(* Logix 5000 project; controller PLC_MCC1201_220AP1 vendor 1 type 14 code 164 rev 35.11; software revision 35.00; part 22 of 25 *)
(* tags used below, declared in another part *)
   LEHR_dActualSpeedValue_mm_min : DINT;
   LEHR_dLehrPositionAdvancement : DINT;
   TMP_dDistanceBetweenCut : DINT;
   TMP_xSimulationMode : BOOL;
   DISTANCE : ALIAS FOR N7[1];
   M203DROP_HMR : MAC_DROPCONV_HMR;
   M225 : MAC_EMERGENCYXCUT;
   M225_ALM : MAC_EMERGENCYXCUT_ALM;
   M225_HMR : MAC_EMERGENCYXCUT_HMR;
   M225_HMW : MAC_EMERGENCYXCUT_HMW;
   M225_IN_MOTION : MAC_EMERGENCYXCUT_IN_MOTION;
   M225_M1_DR : AXIS_CIP_DRIVE;
   M225_OUT_MOTION : MAC_EMERGENCYXCUT_OUT_MOTION;
   N54 : DINT[501];
   Status : INT;   // INT tag to retrieve Status value through GSV created during conversion
   TMP_dIndex : DINT;
   Z200_UPS : ZONE_UPS;
(* MainProgram, continued *)

ROUTINE M225_EmCut_Faults   (* ladder *)
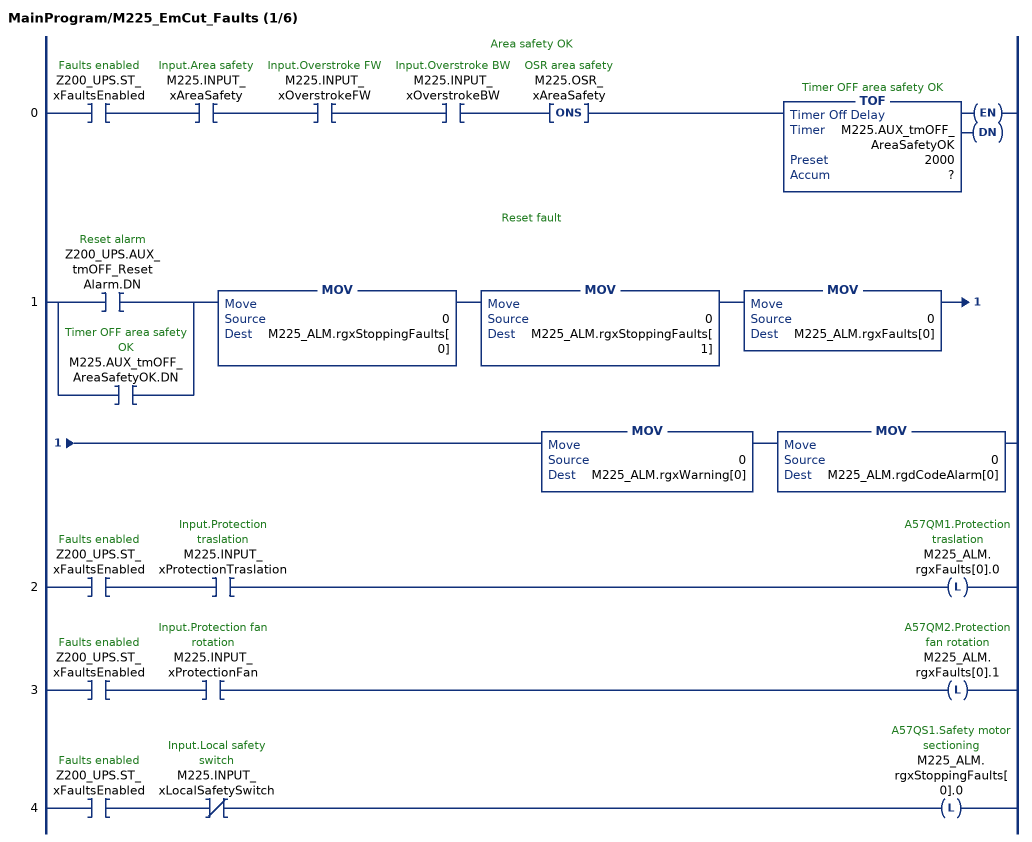
   // Area safety OK
   0: XIC(Z200_UPS.ST_xFaultsEnabled)XIC(M225.INPUT_xAreaSafety)XIC(M225.INPUT_xOverstrokeFW)XIC(M225.INPUT_xOverstrokeBW)ONS(M225.OSR_xAreaSafety)TOF(M225.AUX_tmOFF_AreaSafetyOK,?,?);
   // Reset fault
   1: [XIC(Z200_UPS.AUX_tmOFF_ResetAlarm.DN) ,XIC(M225.AUX_tmOFF_AreaSafetyOK.DN) ]MOV(0,M225_ALM.rgxStoppingFaults[0])MOV(0,M225_ALM.rgxStoppingFaults[1])MOV(0,M225_ALM.rgxFaults[0])MOV(0,M225_ALM.rgxWarning[0])MOV(0,M225_ALM.rgdCodeAlarm[0]);
   2: XIC(Z200_UPS.ST_xFaultsEnabled)XIC(M225.INPUT_xProtectionTraslation)OTL(M225_ALM.rgxFaults[0].0);
   3: XIC(Z200_UPS.ST_xFaultsEnabled)XIC(M225.INPUT_xProtectionFan)OTL(M225_ALM.rgxFaults[0].1);
   4: XIC(Z200_UPS.ST_xFaultsEnabled)XIO(M225.INPUT_xLocalSafetySwitch)OTL(M225_ALM.rgxStoppingFaults[0].0);
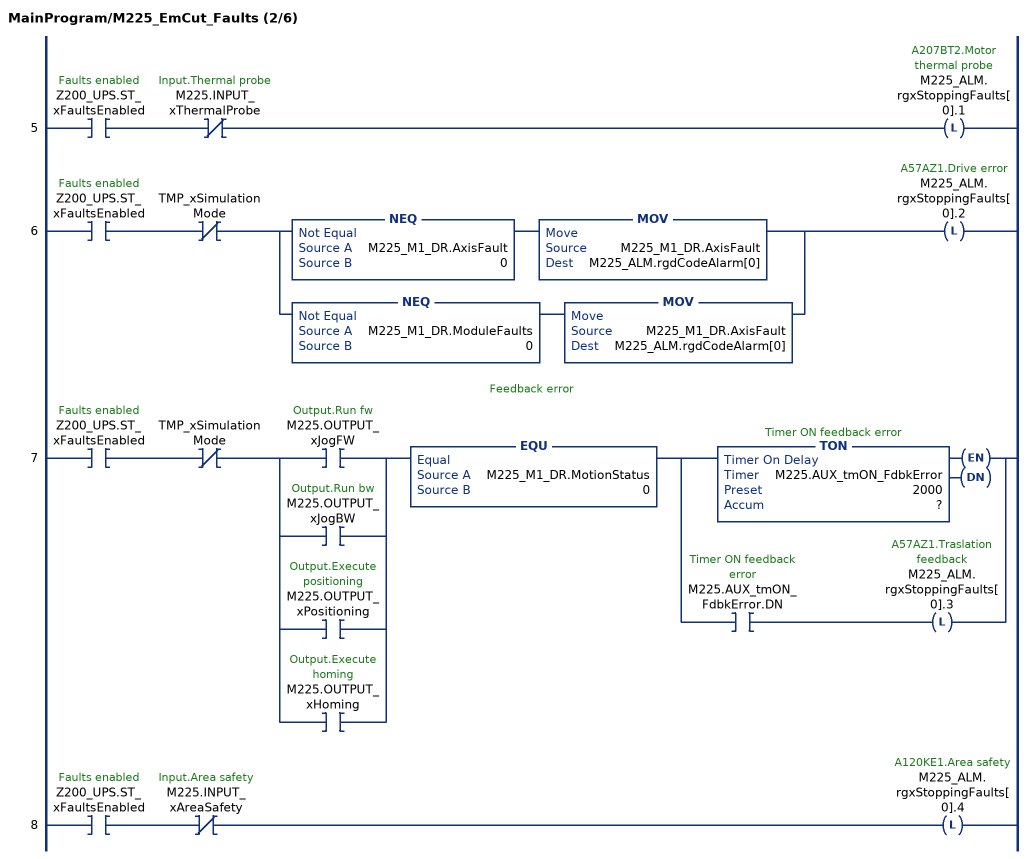
   5: XIC(Z200_UPS.ST_xFaultsEnabled)XIO(M225.INPUT_xThermalProbe)OTL(M225_ALM.rgxStoppingFaults[0].1);
   6: XIC(Z200_UPS.ST_xFaultsEnabled)XIO(TMP_xSimulationMode)[NEQ(M225_M1_DR.AxisFault,0) MOV(M225_M1_DR.AxisFault,M225_ALM.rgdCodeAlarm[0]) ,NEQ(M225_M1_DR.ModuleFaults,0) MOV(M225_M1_DR.AxisFault,M225_ALM.rgdCodeAlarm[0]) ]OTL(M225_ALM.rgxStoppingFaults[0].2);
   // Feedback error
   7: XIC(Z200_UPS.ST_xFaultsEnabled)XIO(TMP_xSimulationMode)[XIC(M225.OUTPUT_xJogFW) ,XIC(M225.OUTPUT_xJogBW) ,XIC(M225.OUTPUT_xPositioning) ,XIC(M225.OUTPUT_xHoming) ]EQU(M225_M1_DR.MotionStatus,0)[TON(M225.AUX_tmON_FdbkError,?,?) ,XIC(M225.AUX_tmON_FdbkError.DN) OTL(M225_ALM.rgxStoppingFaults[0].3) ];
   8: XIC(Z200_UPS.ST_xFaultsEnabled)XIO(M225.INPUT_xAreaSafety)OTL(M225_ALM.rgxStoppingFaults[0].4);
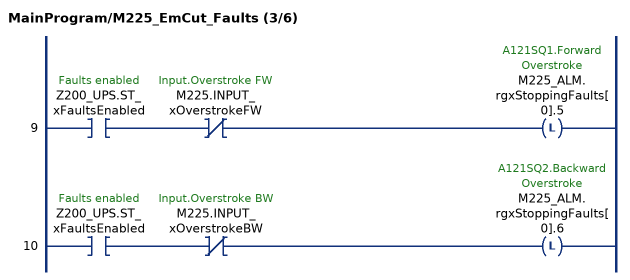
   9: XIC(Z200_UPS.ST_xFaultsEnabled)XIO(M225.INPUT_xOverstrokeFW)OTL(M225_ALM.rgxStoppingFaults[0].5);
   10: XIC(Z200_UPS.ST_xFaultsEnabled)XIO(M225.INPUT_xOverstrokeBW)OTL(M225_ALM.rgxStoppingFaults[0].6);
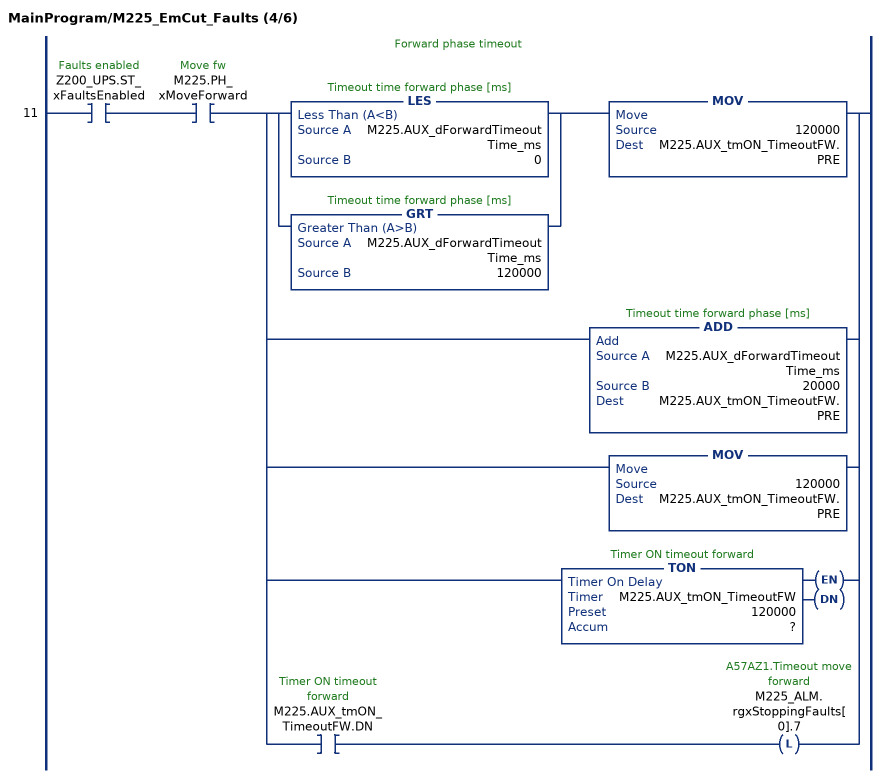
   // Forward phase timeout
   11: XIC(Z200_UPS.ST_xFaultsEnabled)XIC(M225.PH_xMoveForward)[[LES(M225.AUX_dForwardTimeoutTime_ms,0) ,GRT(M225.AUX_dForwardTimeoutTime_ms,120000) ] MOV(120000,M225.AUX_tmON_TimeoutFW.PRE) ,ADD(M225.AUX_dForwardTimeoutTime_ms,20000,M225.AUX_tmON_TimeoutFW.PRE) ,MOV(120000,M225.AUX_tmON_TimeoutFW.PRE) ,TON(M225.AUX_tmON_TimeoutFW,?,?) ,XIC(M225.AUX_tmON_TimeoutFW.DN) OTL(M225_ALM.rgxStoppingFaults[0].7) ];
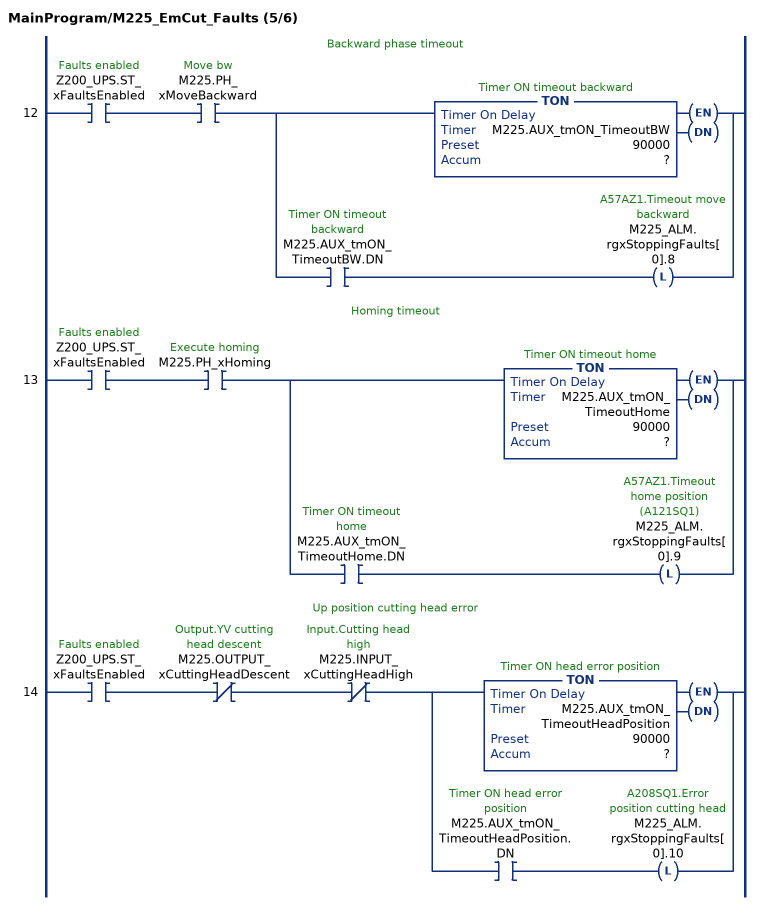
   // Backward phase timeout
   12: XIC(Z200_UPS.ST_xFaultsEnabled)XIC(M225.PH_xMoveBackward)[TON(M225.AUX_tmON_TimeoutBW,?,?) ,XIC(M225.AUX_tmON_TimeoutBW.DN) OTL(M225_ALM.rgxStoppingFaults[0].8) ];
   // Homing timeout
   13: XIC(Z200_UPS.ST_xFaultsEnabled)XIC(M225.PH_xHoming)[TON(M225.AUX_tmON_TimeoutHome,?,?) ,XIC(M225.AUX_tmON_TimeoutHome.DN) OTL(M225_ALM.rgxStoppingFaults[0].9) ];
   // Up position cutting head error
   14: XIC(Z200_UPS.ST_xFaultsEnabled)XIO(M225.OUTPUT_xCuttingHeadDescent)XIO(M225.INPUT_xCuttingHeadHigh)[TON(M225.AUX_tmON_TimeoutHeadPosition,?,?) ,XIC(M225.AUX_tmON_TimeoutHeadPosition.DN) OTL(M225_ALM.rgxStoppingFaults[0].10) ];
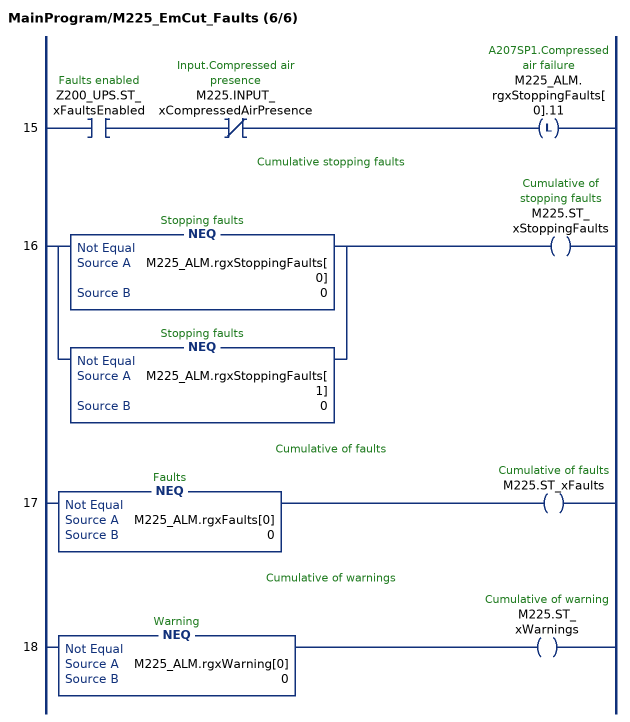
   15: XIC(Z200_UPS.ST_xFaultsEnabled)XIO(M225.INPUT_xCompressedAirPresence)OTL(M225_ALM.rgxStoppingFaults[0].11);
   // Cumulative stopping faults
   16: [NEQ(M225_ALM.rgxStoppingFaults[0],0) ,NEQ(M225_ALM.rgxStoppingFaults[1],0) ]OTE(M225.ST_xStoppingFaults);
   // Cumulative of faults
   17: NEQ(M225_ALM.rgxFaults[0],0)OTE(M225.ST_xFaults);
   // Cumulative of warnings
   18: NEQ(M225_ALM.rgxWarning[0],0)OTE(M225.ST_xWarnings);
END_ROUTINE

ROUTINE M225_EmCut_FIFOTank   (* structured text *)
   FOR TMP_dIndex:=0 TO M225.AUX_dTankElementCounter-1 DO
   	M225.AUX_rgdCutTank[TMP_dIndex]:=M225.AUX_rgdCutTank[TMP_dIndex+1];
   END_FOR;
END_ROUTINE

ROUTINE M225_EmCut_Logics   (* ladder *)
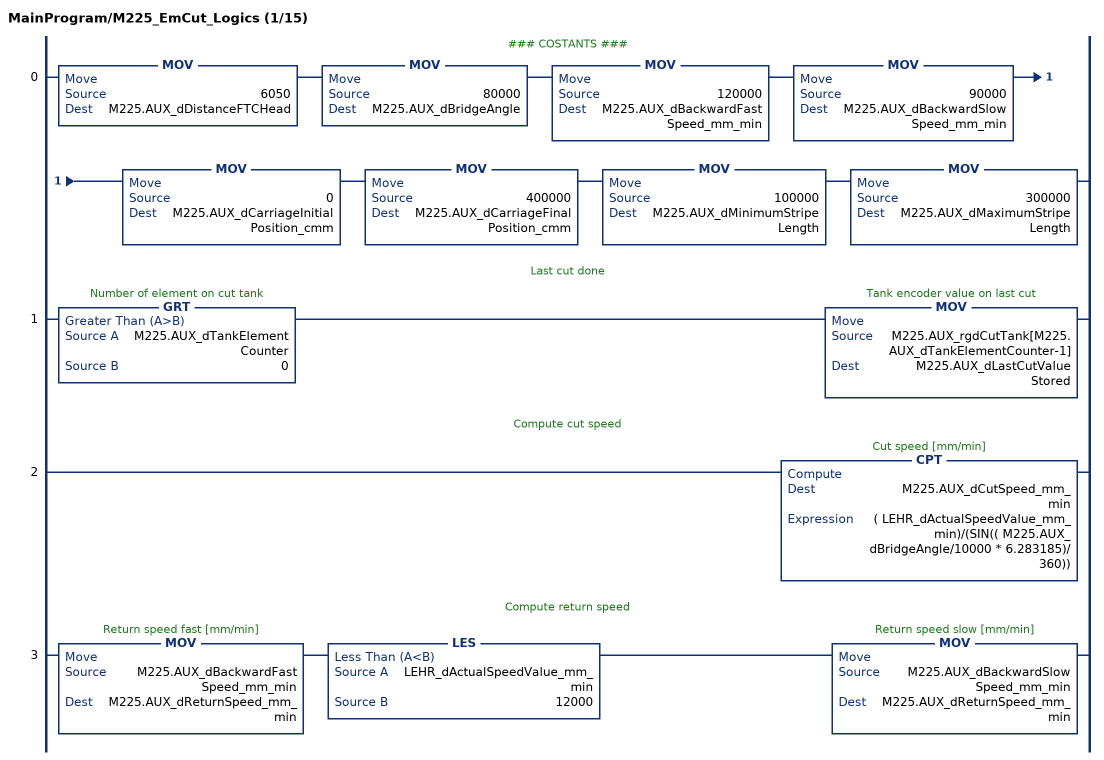
   // ### COSTANTS ###
   0: MOV(6050,M225.AUX_dDistanceFTCHead)MOV(80000,M225.AUX_dBridgeAngle)MOV(120000,M225.AUX_dBackwardFastSpeed_mm_min)MOV(90000,M225.AUX_dBackwardSlowSpeed_mm_min)MOV(0,M225.AUX_dCarriageInitialPosition_cmm)MOV(400000,M225.AUX_dCarriageFinalPosition_cmm)MOV(100000,M225.AUX_dMinimumStripeLength)MOV(300000,M225.AUX_dMaximumStripeLength);
   // Last cut done
   1: GRT(M225.AUX_dTankElementCounter,0)MOV(M225.AUX_rgdCutTank[M225.AUX_dTankElementCounter-1],M225.AUX_dLastCutValueStored);
   // Compute cut speed
   2: CPT(M225.AUX_dCutSpeed_mm_min,( LEHR_dActualSpeedValue_mm_min)/(SIN(( M225.AUX_dBridgeAngle/10000 * 6.283185)/ 360)));
   // Compute return speed
   3: MOV(M225.AUX_dBackwardFastSpeed_mm_min,M225.AUX_dReturnSpeed_mm_min)LES(LEHR_dActualSpeedValue_mm_min,12000)MOV(M225.AUX_dBackwardSlowSpeed_mm_min,M225.AUX_dReturnSpeed_mm_min);
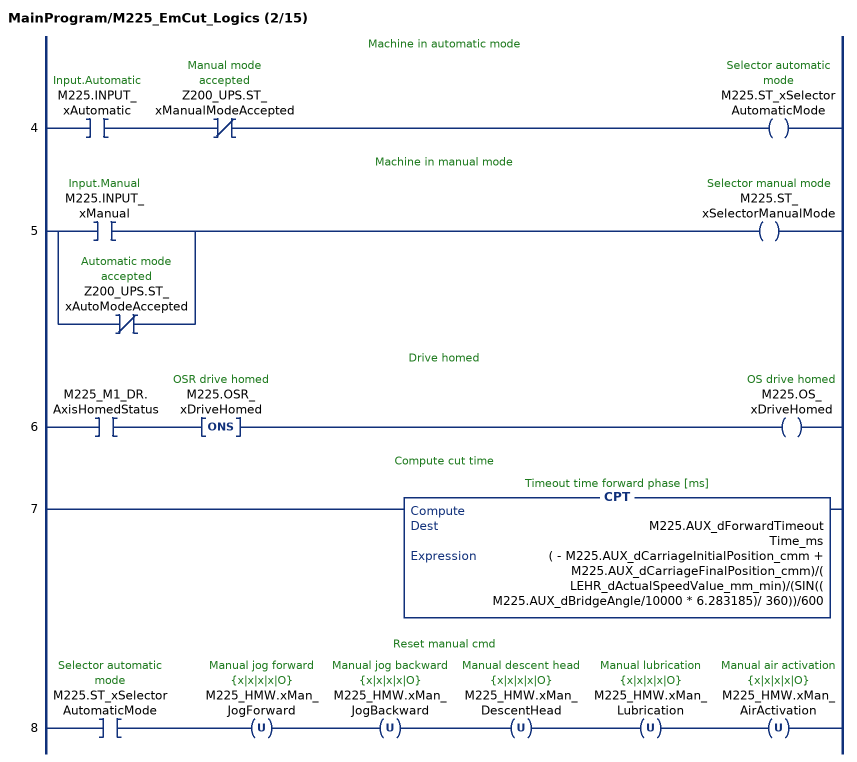
   // Machine in automatic mode
   4: XIC(M225.INPUT_xAutomatic)XIO(Z200_UPS.ST_xManualModeAccepted)OTE(M225.ST_xSelectorAutomaticMode);
   // Machine in manual mode
   5: [XIC(M225.INPUT_xManual) ,XIO(Z200_UPS.ST_xAutoModeAccepted) ]OTE(M225.ST_xSelectorManualMode);
   // Drive homed
   6: XIC(M225_M1_DR.AxisHomedStatus)ONS(M225.OSR_xDriveHomed)OTE(M225.OS_xDriveHomed);
   // Compute cut time
   7: CPT(M225.AUX_dForwardTimeoutTime_ms,( - M225.AUX_dCarriageInitialPosition_cmm + M225.AUX_dCarriageFinalPosition_cmm)/( LEHR_dActualSpeedValue_mm_min)/(SIN(( M225.AUX_dBridgeAngle/10000 * 6.283185)/ 360))/600);
   // Reset manual cmd
   8: XIC(M225.ST_xSelectorAutomaticMode)OTU(M225_HMW.xMan_JogForward)OTU(M225_HMW.xMan_JogBackward)OTU(M225_HMW.xMan_DescentHead)OTU(M225_HMW.xMan_Lubrication)OTU(M225_HMW.xMan_AirActivation);
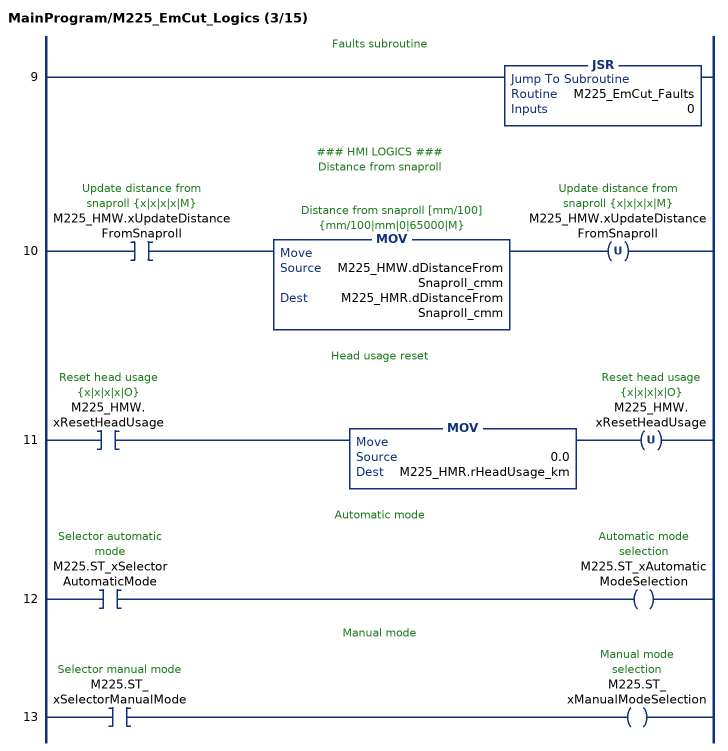
   // Faults subroutine
   9: JSR(M225_EmCut_Faults,0);
   // ### HMI LOGICS ###
   // Distance from snaproll
   10: XIC(M225_HMW.xUpdateDistanceFromSnaproll)MOV(M225_HMW.dDistanceFromSnaproll_cmm,M225_HMR.dDistanceFromSnaproll_cmm)OTU(M225_HMW.xUpdateDistanceFromSnaproll);
   // Head usage reset
   11: XIC(M225_HMW.xResetHeadUsage)MOV(0.0,M225_HMR.rHeadUsage_km)OTU(M225_HMW.xResetHeadUsage);
   // Automatic mode
   12: XIC(M225.ST_xSelectorAutomaticMode)OTE(M225.ST_xAutomaticModeSelection);
   // Manual mode
   13: XIC(M225.ST_xSelectorManualMode)OTE(M225.ST_xManualModeSelection);
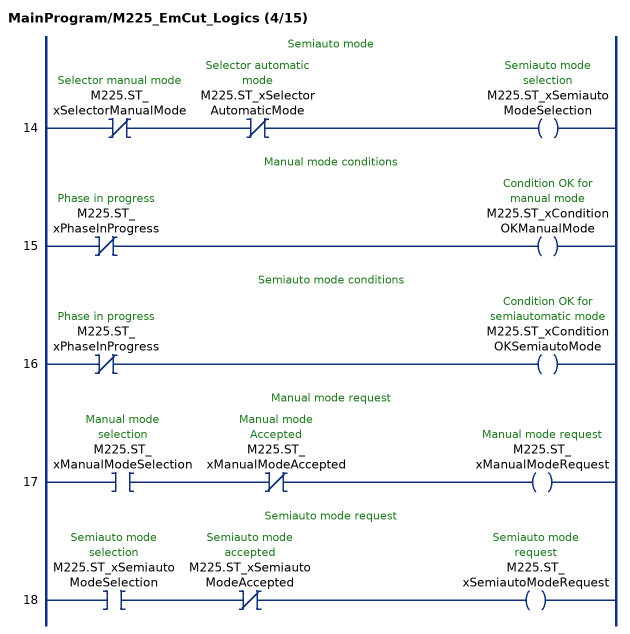
   // Semiauto mode
   14: XIO(M225.ST_xSelectorManualMode)XIO(M225.ST_xSelectorAutomaticMode)OTE(M225.ST_xSemiautoModeSelection);
   // Manual mode conditions
   15: XIO(M225.ST_xPhaseInProgress)OTE(M225.ST_xConditionOKManualMode);
   // Semiauto mode conditions
   16: XIO(M225.ST_xPhaseInProgress)OTE(M225.ST_xConditionOKSemiautoMode);
   // Manual mode request
   17: XIC(M225.ST_xManualModeSelection)XIO(M225.ST_xManualModeAccepted)OTE(M225.ST_xManualModeRequest);
   // Semiauto mode request
   18: XIC(M225.ST_xSemiautoModeSelection)XIO(M225.ST_xSemiautoModeAccepted)OTE(M225.ST_xSemiautoModeRequest);
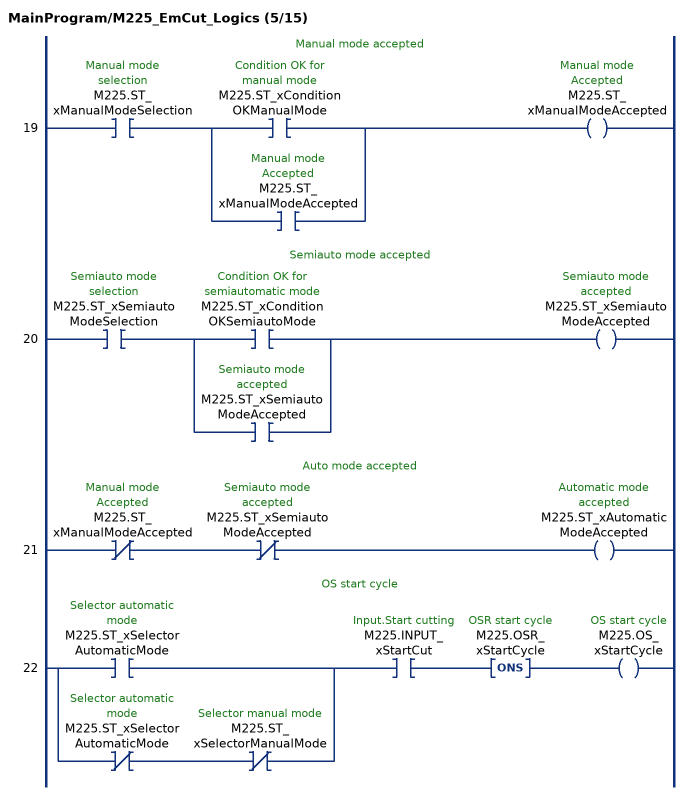
   // Manual mode accepted
   19: XIC(M225.ST_xManualModeSelection)[XIC(M225.ST_xConditionOKManualMode) ,XIC(M225.ST_xManualModeAccepted) ]OTE(M225.ST_xManualModeAccepted);
   // Semiauto mode accepted
   20: XIC(M225.ST_xSemiautoModeSelection)[XIC(M225.ST_xConditionOKSemiautoMode) ,XIC(M225.ST_xSemiautoModeAccepted) ]OTE(M225.ST_xSemiautoModeAccepted);
   // Auto mode accepted
   21: XIO(M225.ST_xManualModeAccepted)XIO(M225.ST_xSemiautoModeAccepted)OTE(M225.ST_xAutomaticModeAccepted);
   // OS start cycle
   22: [XIC(M225.ST_xSelectorAutomaticMode) ,XIO(M225.ST_xSelectorAutomaticMode) XIO(M225.ST_xSelectorManualMode) ]XIC(M225.INPUT_xStartCut)ONS(M225.OSR_xStartCycle)OTE(M225.OS_xStartCycle);
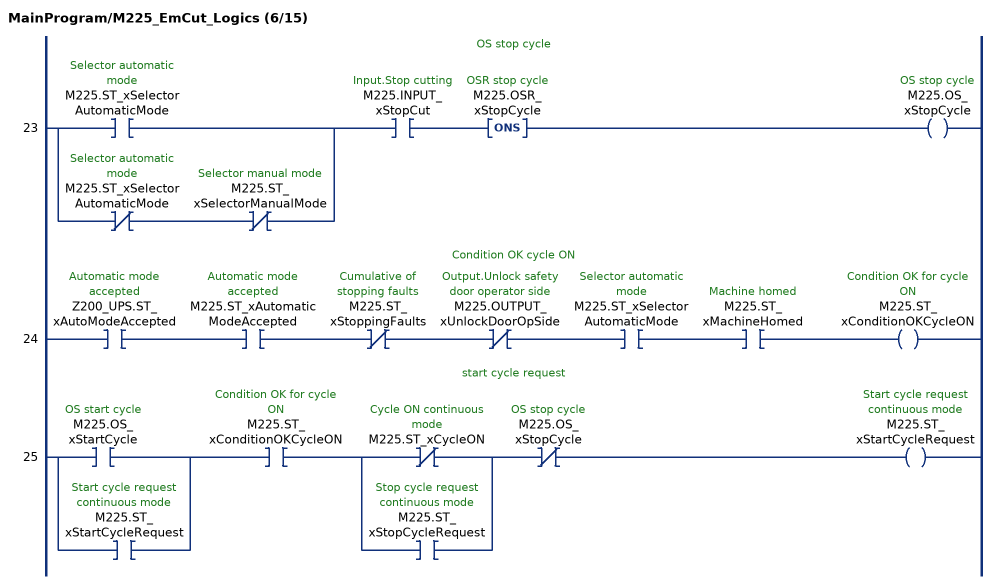
   // OS stop cycle
   23: [XIC(M225.ST_xSelectorAutomaticMode) ,XIO(M225.ST_xSelectorAutomaticMode) XIO(M225.ST_xSelectorManualMode) ]XIC(M225.INPUT_xStopCut)ONS(M225.OSR_xStopCycle)OTE(M225.OS_xStopCycle);
   // Condition OK cycle ON
   24: XIC(Z200_UPS.ST_xAutoModeAccepted)XIC(M225.ST_xAutomaticModeAccepted)XIO(M225.ST_xStoppingFaults)XIO(M225.OUTPUT_xUnlockDoorOpSide)XIC(M225.ST_xSelectorAutomaticMode)XIC(M225.ST_xMachineHomed)OTE(M225.ST_xConditionOKCycleON);
   // start cycle request
   25: [XIC(M225.OS_xStartCycle) ,XIC(M225.ST_xStartCycleRequest) ]XIC(M225.ST_xConditionOKCycleON)[XIO(M225.ST_xCycleON) ,XIC(M225.ST_xStopCycleRequest) ]XIO(M225.OS_xStopCycle)OTE(M225.ST_xStartCycleRequest);
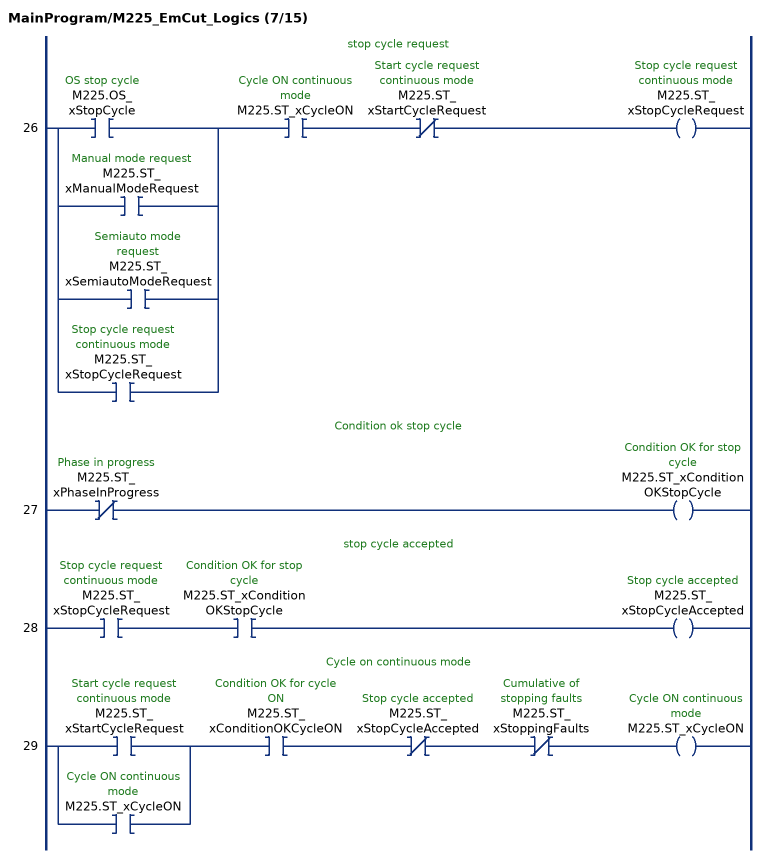
   // stop cycle request
   26: [XIC(M225.OS_xStopCycle) ,XIC(M225.ST_xManualModeRequest) ,XIC(M225.ST_xSemiautoModeRequest) ,XIC(M225.ST_xStopCycleRequest) ]XIC(M225.ST_xCycleON)XIO(M225.ST_xStartCycleRequest)OTE(M225.ST_xStopCycleRequest);
   // Condition ok stop cycle
   27: XIO(M225.ST_xPhaseInProgress)OTE(M225.ST_xConditionOKStopCycle);
   // stop cycle accepted
   28: XIC(M225.ST_xStopCycleRequest)XIC(M225.ST_xConditionOKStopCycle)OTE(M225.ST_xStopCycleAccepted);
   // Cycle on continuous mode
   29: [XIC(M225.ST_xStartCycleRequest) ,XIC(M225.ST_xCycleON) ]XIC(M225.ST_xConditionOKCycleON)XIO(M225.ST_xStopCycleAccepted)XIO(M225.ST_xStoppingFaults)OTE(M225.ST_xCycleON);
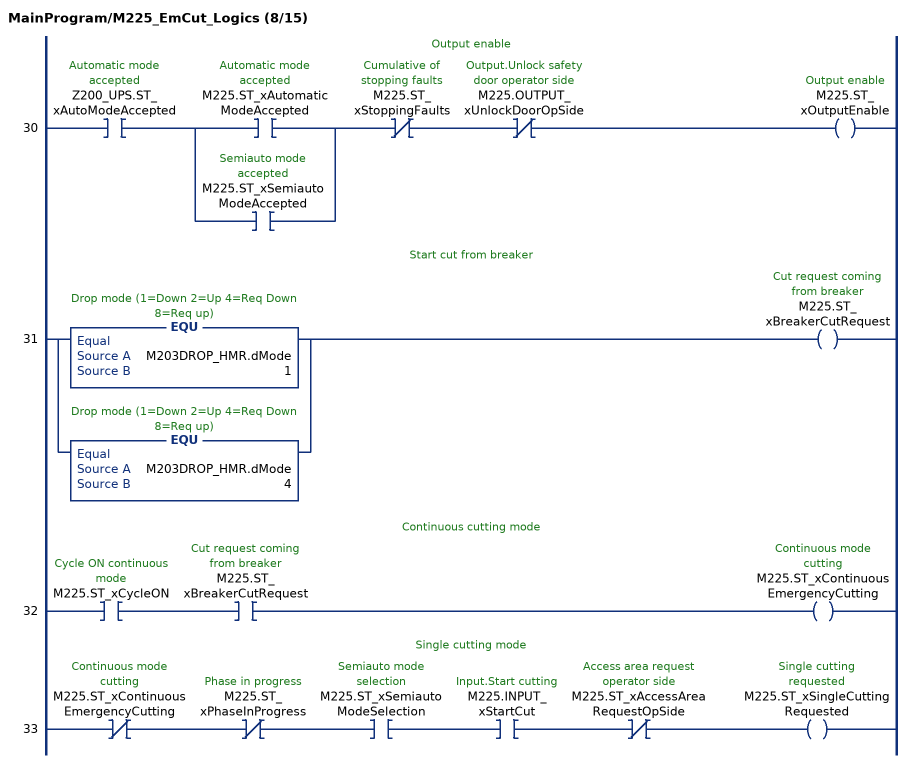
   // Output enable
   30: XIC(Z200_UPS.ST_xAutoModeAccepted)[XIC(M225.ST_xAutomaticModeAccepted) ,XIC(M225.ST_xSemiautoModeAccepted) ]XIO(M225.ST_xStoppingFaults)XIO(M225.OUTPUT_xUnlockDoorOpSide)OTE(M225.ST_xOutputEnable);
   // Start cut from breaker
   31: [EQU(M203DROP_HMR.dMode,1) ,EQU(M203DROP_HMR.dMode,4) ]OTE(M225.ST_xBreakerCutRequest);
   // Continuous cutting mode
   32: XIC(M225.ST_xCycleON)XIC(M225.ST_xBreakerCutRequest)OTE(M225.ST_xContinuousEmergencyCutting);
   // Single cutting mode
   33: XIO(M225.ST_xContinuousEmergencyCutting)XIO(M225.ST_xPhaseInProgress)XIC(M225.ST_xSemiautoModeSelection)XIC(M225.INPUT_xStartCut)XIO(M225.ST_xAccessAreaRequestOpSide)OTE(M225.ST_xSingleCuttingRequested);
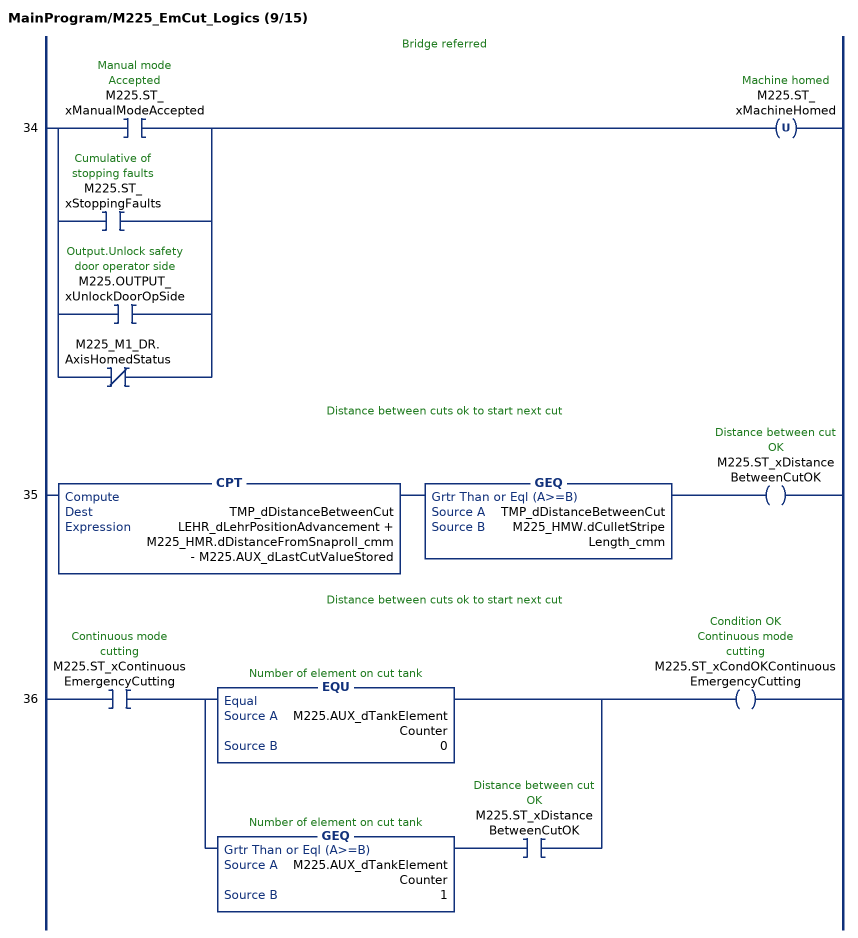
   // Bridge referred
   34: [XIC(M225.ST_xManualModeAccepted) ,XIC(M225.ST_xStoppingFaults) ,XIC(M225.OUTPUT_xUnlockDoorOpSide) ,XIO(M225_M1_DR.AxisHomedStatus) ]OTU(M225.ST_xMachineHomed);
   // Distance between cuts ok to start next cut
   35: CPT(TMP_dDistanceBetweenCut,LEHR_dLehrPositionAdvancement + M225_HMR.dDistanceFromSnaproll_cmm - M225.AUX_dLastCutValueStored)GEQ(TMP_dDistanceBetweenCut,M225_HMW.dCulletStripeLength_cmm)OTE(M225.ST_xDistanceBetweenCutOK);
   // Distance between cuts ok to start next cut
   36: XIC(M225.ST_xContinuousEmergencyCutting)[EQU(M225.AUX_dTankElementCounter,0) ,GEQ(M225.AUX_dTankElementCounter,1) XIC(M225.ST_xDistanceBetweenCutOK) ]OTE(M225.ST_xCondOKContinuousEmergencyCutting);
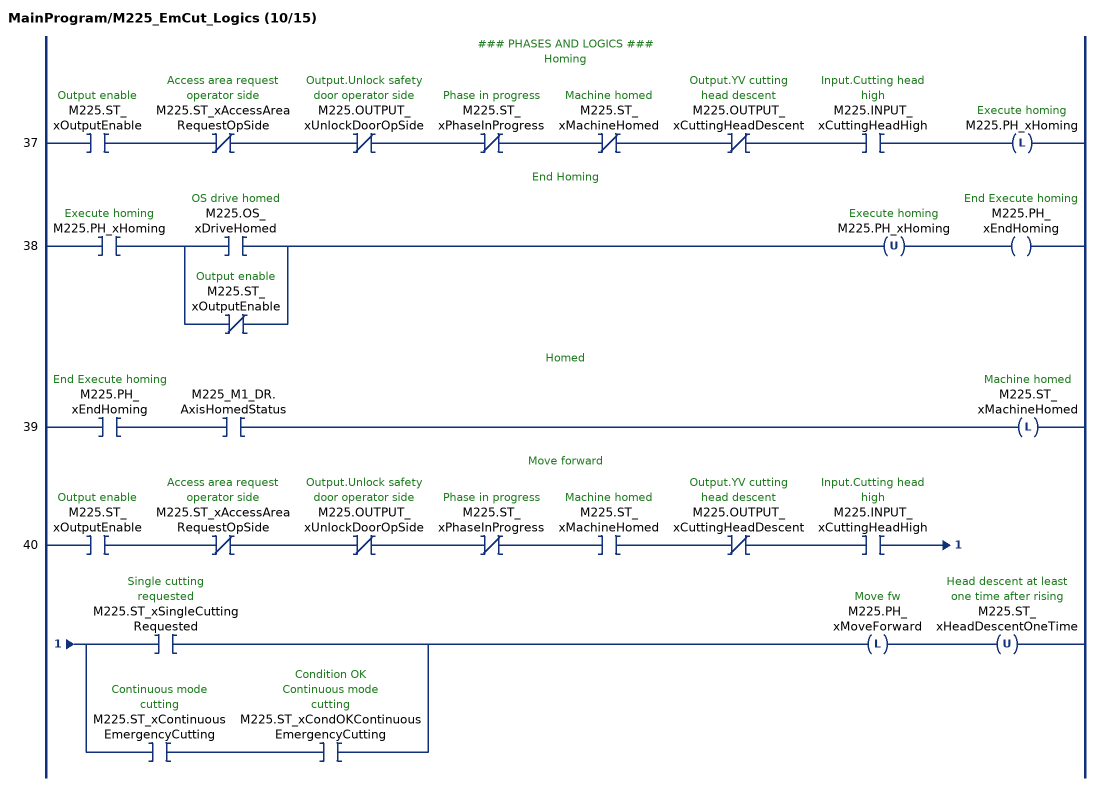
   // ### PHASES AND LOGICS ###
   // Homing
   37: XIC(M225.ST_xOutputEnable)XIO(M225.ST_xAccessAreaRequestOpSide)XIO(M225.OUTPUT_xUnlockDoorOpSide)XIO(M225.ST_xPhaseInProgress)XIO(M225.ST_xMachineHomed)XIO(M225.OUTPUT_xCuttingHeadDescent)XIC(M225.INPUT_xCuttingHeadHigh)OTL(M225.PH_xHoming);
   // End Homing
   38: XIC(M225.PH_xHoming)[XIC(M225.OS_xDriveHomed) ,XIO(M225.ST_xOutputEnable) ]OTU(M225.PH_xHoming)OTE(M225.PH_xEndHoming);
   // Homed
   39: XIC(M225.PH_xEndHoming)XIC(M225_M1_DR.AxisHomedStatus)OTL(M225.ST_xMachineHomed);
   // Move forward
   40: XIC(M225.ST_xOutputEnable)XIO(M225.ST_xAccessAreaRequestOpSide)XIO(M225.OUTPUT_xUnlockDoorOpSide)XIO(M225.ST_xPhaseInProgress)XIC(M225.ST_xMachineHomed)XIO(M225.OUTPUT_xCuttingHeadDescent)XIC(M225.INPUT_xCuttingHeadHigh)[XIC(M225.ST_xSingleCuttingRequested) ,XIC(M225.ST_xContinuousEmergencyCutting) XIC(M225.ST_xCondOKContinuousEmergencyCutting) ]OTL(M225.PH_xMoveForward)OTU(M225.ST_xHeadDescentOneTime);
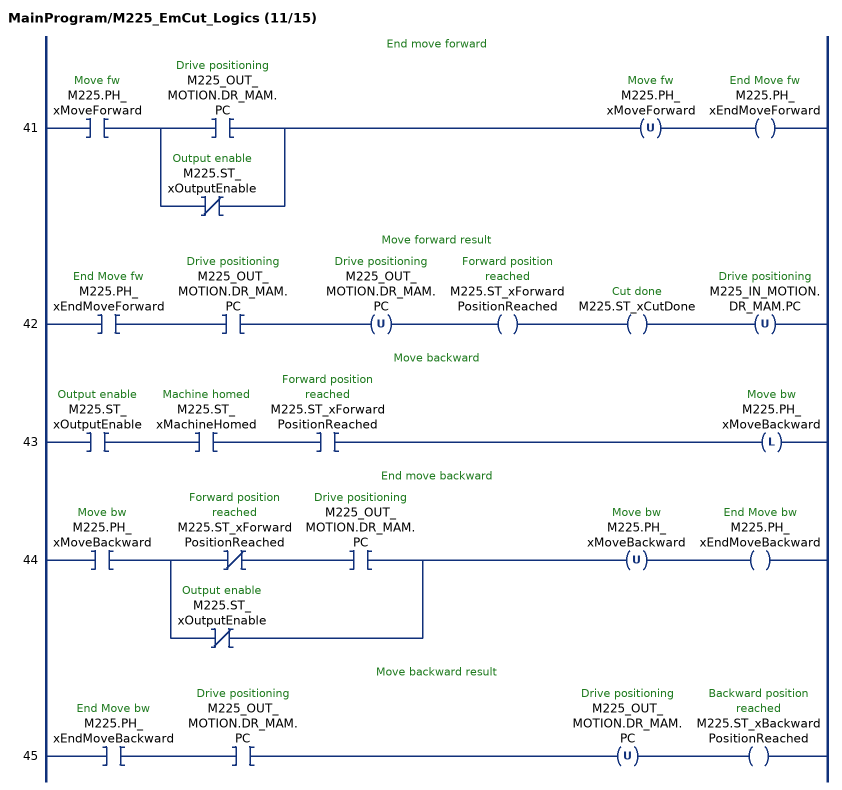
   // End move forward
   41: XIC(M225.PH_xMoveForward)[XIC(M225_OUT_MOTION.DR_MAM.PC) ,XIO(M225.ST_xOutputEnable) ]OTU(M225.PH_xMoveForward)OTE(M225.PH_xEndMoveForward);
   // Move forward result
   42: XIC(M225.PH_xEndMoveForward)XIC(M225_OUT_MOTION.DR_MAM.PC)OTU(M225_OUT_MOTION.DR_MAM.PC)OTE(M225.ST_xForwardPositionReached)OTE(M225.ST_xCutDone)OTU(M225_IN_MOTION.DR_MAM.PC);
   // Move backward
   43: XIC(M225.ST_xOutputEnable)XIC(M225.ST_xMachineHomed)XIC(M225.ST_xForwardPositionReached)OTL(M225.PH_xMoveBackward);
   // End move backward
   44: XIC(M225.PH_xMoveBackward)[XIO(M225.ST_xForwardPositionReached) XIC(M225_OUT_MOTION.DR_MAM.PC) ,XIO(M225.ST_xOutputEnable) ]OTU(M225.PH_xMoveBackward)OTE(M225.PH_xEndMoveBackward);
   // Move backward result
   45: XIC(M225.PH_xEndMoveBackward)XIC(M225_OUT_MOTION.DR_MAM.PC)OTU(M225_OUT_MOTION.DR_MAM.PC)OTE(M225.ST_xBackwardPositionReached);
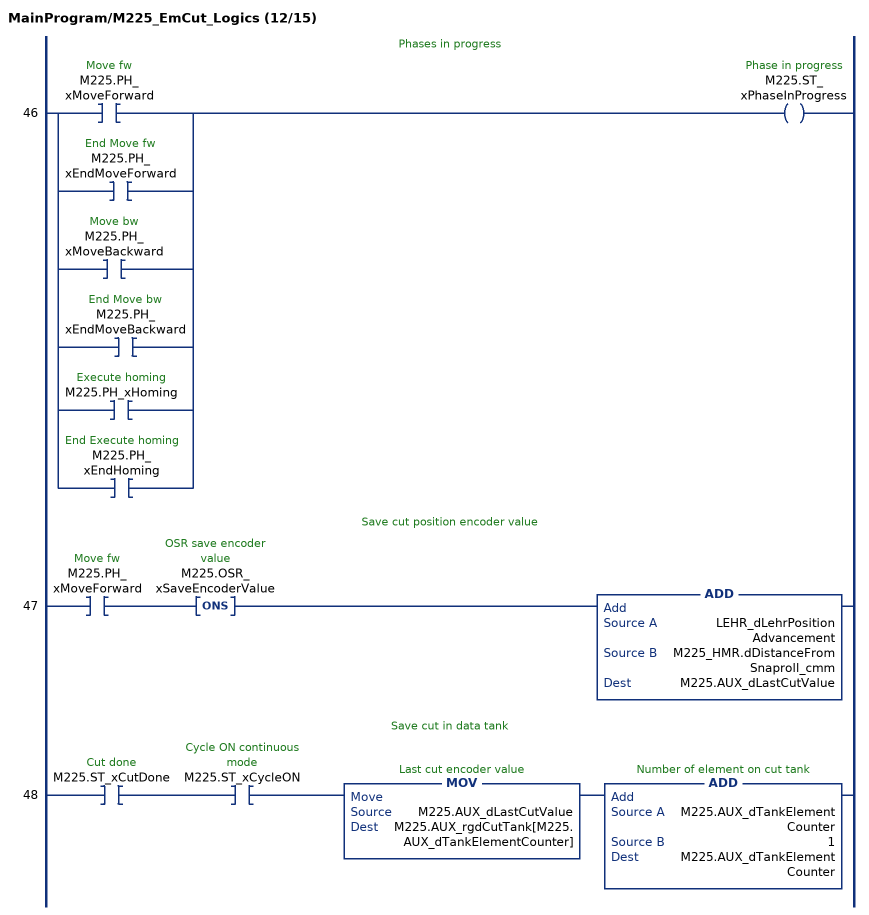
   // Phases in progress
   46: [XIC(M225.PH_xMoveForward) ,XIC(M225.PH_xEndMoveForward) ,XIC(M225.PH_xMoveBackward) ,XIC(M225.PH_xEndMoveBackward) ,XIC(M225.PH_xHoming) ,XIC(M225.PH_xEndHoming) ]OTE(M225.ST_xPhaseInProgress);
   // Save cut position encoder value
   47: XIC(M225.PH_xMoveForward)ONS(M225.OSR_xSaveEncoderValue)ADD(LEHR_dLehrPositionAdvancement,M225_HMR.dDistanceFromSnaproll_cmm,M225.AUX_dLastCutValue);
   // Save cut in data tank
   48: XIC(M225.ST_xCutDone)XIC(M225.ST_xCycleON)MOV(M225.AUX_dLastCutValue,M225.AUX_rgdCutTank[M225.AUX_dTankElementCounter])ADD(M225.AUX_dTankElementCounter,1,M225.AUX_dTankElementCounter);
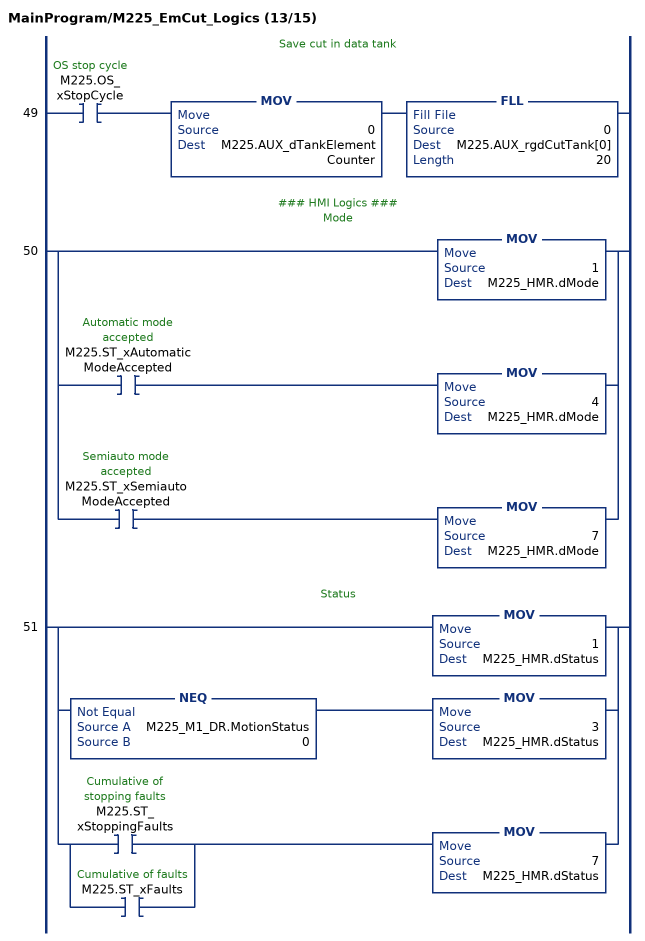
   // Save cut in data tank
   49: XIC(M225.OS_xStopCycle)MOV(0,M225.AUX_dTankElementCounter)FLL(0,M225.AUX_rgdCutTank[0],20);
   // ### HMI Logics ###
   // Mode
   50: [MOV(1,M225_HMR.dMode) ,XIC(M225.ST_xAutomaticModeAccepted) MOV(4,M225_HMR.dMode) ,XIC(M225.ST_xSemiautoModeAccepted) MOV(7,M225_HMR.dMode) ];
   // Status
   51: [MOV(1,M225_HMR.dStatus) ,NEQ(M225_M1_DR.MotionStatus,0) MOV(3,M225_HMR.dStatus) ,[XIC(M225.ST_xStoppingFaults) ,XIC(M225.ST_xFaults) ] MOV(7,M225_HMR.dStatus) ];
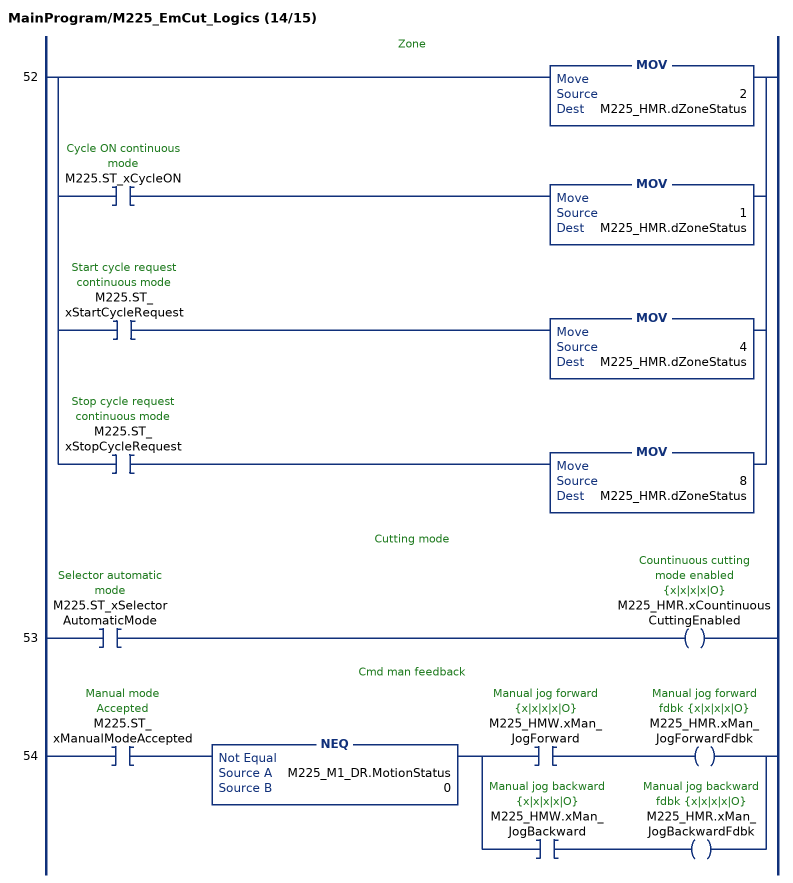
   // Zone
   52: [MOV(2,M225_HMR.dZoneStatus) ,XIC(M225.ST_xCycleON) MOV(1,M225_HMR.dZoneStatus) ,XIC(M225.ST_xStartCycleRequest) MOV(4,M225_HMR.dZoneStatus) ,XIC(M225.ST_xStopCycleRequest) MOV(8,M225_HMR.dZoneStatus) ];
   // Cutting mode
   53: XIC(M225.ST_xSelectorAutomaticMode)OTE(M225_HMR.xCountinuousCuttingEnabled);
   // Cmd man feedback
   54: XIC(M225.ST_xManualModeAccepted)NEQ(M225_M1_DR.MotionStatus,0)[XIC(M225_HMW.xMan_JogForward) OTE(M225_HMR.xMan_JogForwardFdbk) ,XIC(M225_HMW.xMan_JogBackward) OTE(M225_HMR.xMan_JogBackwardFdbk) ];
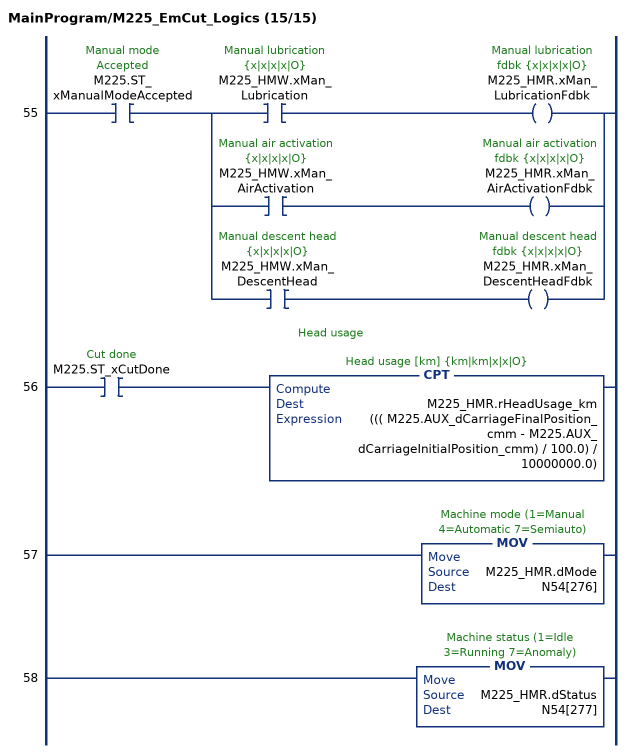
   55: XIC(M225.ST_xManualModeAccepted)[XIC(M225_HMW.xMan_Lubrication) OTE(M225_HMR.xMan_LubricationFdbk) ,XIC(M225_HMW.xMan_AirActivation) OTE(M225_HMR.xMan_AirActivationFdbk) ,XIC(M225_HMW.xMan_DescentHead) OTE(M225_HMR.xMan_DescentHeadFdbk) ];
   // Head usage
   56: XIC(M225.ST_xCutDone)CPT(M225_HMR.rHeadUsage_km,((( M225.AUX_dCarriageFinalPosition_cmm - M225.AUX_dCarriageInitialPosition_cmm) / 100.0) / 10000000.0));
   57: MOV(M225_HMR.dMode,N54[276]);
   58: MOV(M225_HMR.dStatus,N54[277]);
END_ROUTINE
